// TIA Portal project "Project2_Pompe" (V15.1)

(* hardware
DEVICE "S71500/ET200MP station_1"  S7-1500 station
   slot 0: "Rail_0"  Rack  6ES7 590-1***0-0AA0
   slot 1: "PLC_1"  CPU 1513-1 PN  6ES7 513-1AL02-0AB0  V2.6
      slot 3: "CPU display_1"  6ES7591-1AA00-0AA0
DEVICE "HMI_1"  KTP900 Basic PN
   slot 0: "HMI_1"  KTP900 Basic PN  6AV2 123-2JB03-0AX0  15.1.0.0
   slot 1: "HMI_RT_1"  KTP900 Basic PN  6AV2 123-2JB03-0AX0  15.1.0.0
   slot 5: "HMI_1.IE_CP_1"  PROFINET Interface  15.0.1.0
      slot 1: "PROFINET Interface_1"  PROFINET Interface
         slot 1: "Port_1"  Port
*)

// ===== PLC "PLC_1"  CPU 1513-1 PN =====

VAR_GLOBAL   // PLC tag table "Default tag table"
   "Clock_Byte" AT %MB0 : Byte;
   "Clock_10Hz" AT %M0.0 : Bool;
   "Clock_5Hz" AT %M0.1 : Bool;
   "Clock_2.5Hz" AT %M0.2 : Bool;
   "Clock_2Hz" AT %M0.3 : Bool;
   "Clock_1.25Hz" AT %M0.4 : Bool;
   "Clock_1Hz" AT %M0.5 : Bool;
   "Clock_0.625Hz" AT %M0.6 : Bool;
   "Clock_0.5Hz" AT %M0.7 : Bool;
END_VAR

VAR_GLOBAL   // PLC tag table "Motor1"
   "permisie_start_1" AT %I0.0 : Bool;
   "motor_pornit_1" AT %I0.1 : Bool;
   "temporizare_k4_1" AT %I0.2 : Bool;
   "urgenta_bit_1" AT %I0.4 : Bool;
   "s1_1" AT %I0.7 : Bool;
   "s2_1" AT %I1.0 : Bool;
   "stop1" AT %I1.1 : Bool;
   "ptc1" AT %I1.2 : Bool;
   "timp_oprire_1" AT %ID1 : Time;
   "k1_1" AT %M1.4 : Bool;
   "k2_1" AT %M1.5 : Bool;
   "k3_1" AT %M1.6 : Bool;
   "k4_1" AT %M1.7 : Bool;
   "reset_urgenta_1" AT %I7.0 : Bool;
   "et_k4_1" AT %ID11 : Time;
   "et_stop_1" AT %ID10 : Time;
   "inactiv_1" AT %ID20 : Time;
END_VAR

VAR_GLOBAL   // PLC tag table "Motor2"
   "permisie_start_2" AT %I2.0 : Bool;
   "motor_pornit_2" AT %I2.1 : Bool;
   "temporizare_k4_2" AT %I2.2 : Bool;
   "urgenta_bit_2" AT %I2.3 : Bool;
   "s1_2" AT %I2.4 : Bool;
   "s2_2" AT %I2.5 : Bool;
   "stop2" AT %I2.6 : Bool;
   "ptc2" AT %I2.7 : Bool;
   "timp_oprire_2" AT %ID3 : Time;
   "k1_2" AT %M3.1 : Bool;
   "k2_2" AT %M3.2 : Bool;
   "k3_2" AT %M3.3 : Bool;
   "k4_2" AT %M3.4 : Bool;
   "reset_urgenta_2" AT %I7.1 : Bool;
   "et_k4_2" AT %ID7 : Time;
   "et_stop_2" AT %ID12 : Time;
   "inactiv_2" AT %ID16 : Time;
END_VAR

VAR_GLOBAL   // PLC tag table "Ambele_motoare"
   "ss(esd)" AT %I0.6 : Bool;
   "ptc" AT %I36.0 : Bool;
   "stop" AT %I36.1 : Bool;
   "reset_urgenta_general" AT %I36.2 : Bool;
   "urgenta_bit_ciuperca" AT %I36.3 : Bool;
   "oprire_toate_motoarele_pt_ptc" AT %I36.4 : Bool;
END_VAR

VAR_GLOBAL   // PLC tag table "Motor3"
   "permisie_start_3" AT %I30.0 : Bool;
   "motor_pornit_3" AT %I30.1 : Bool;
   "temporizare_k4_3" AT %I30.2 : Bool;
   "urgenta_bit_3" AT %I30.3 : Bool;
   "s1_3" AT %I30.4 : Bool;
   "s2_3" AT %I30.5 : Bool;
   "stop3" AT %I30.6 : Bool;
   "ptc3" AT %I30.7 : Bool;
   "k1_3" AT %M31.0 : Bool;
   "k2_3" AT %M31.1 : Bool;
   "k3_3" AT %M31.2 : Bool;
   "k4_3" AT %M31.3 : Bool;
   "reset_urgenta_3" AT %I31.4 : Bool;
   "et_k4_3" AT %ID31 : Time;
   "et_stop_3" AT %ID32 : Time;
END_VAR

VAR_GLOBAL   // PLC tag table "Motor4"
   "permisie_start_4" AT %I0.3 : Bool;
   "motor_pornit_4" AT %I0.5 : Bool;
   "temporizare_k4_4" AT %I24.0 : Bool;
   "urgenta_bit_4" AT %I24.1 : Bool;
   "s1_4" AT %I24.2 : Bool;
   "s2_4" AT %I24.3 : Bool;
   "stop4" AT %I24.4 : Bool;
   "pct4" AT %I24.5 : Bool;
   "k1_4" AT %M24.6 : Bool;
   "k2_4" AT %M24.7 : Bool;
   "k3_4" AT %M25.0 : Bool;
   "k4_4" AT %M25.1 : Bool;
   "reset_urgenta_4" AT %I25.2 : Bool;
   "et_k4_4" AT %ID25 : Time;
   "et_stop_4" AT %ID26 : Time;
END_VAR

DATA_BLOCK "db_directie_mers"   // DB1
{ S7_Optimized_Access := 'TRUE' }
VERSION : 0.1
   VAR
      et_stop : Time;
      stanga : Bool;
      dreapta : Bool;
      inainte : Bool;
      inapoi : Bool;
      stop : Bool;
   END_VAR
BEGIN
END_DATA_BLOCK

DATA_BLOCK "roata 2"   // DB3
{ S7_Optimized_Access := 'TRUE' }
VERSION : 0.1
// stored: InstanceOfName Fct_Motor
"Fct_Motor"
BEGIN
END_DATA_BLOCK

DATA_BLOCK "roata 3"   // DB4
{ S7_Optimized_Access := 'TRUE' }
VERSION : 0.1
// stored: InstanceOfName Fct_Motor
"Fct_Motor"
BEGIN
END_DATA_BLOCK

DATA_BLOCK "Alarme"   // DB5
{ S7_Optimized_Access := 'TRUE' }
VERSION : 0.1
   VAR
      alarme : Array[0..15] of Bool;
      alarme_merged : Word;
   END_VAR
BEGIN
END_DATA_BLOCK

DATA_BLOCK "functie ptc_DB_r1"   // DB7
{ S7_Optimized_Access := 'TRUE' }
VERSION : 0.1
// stored: InstanceOfName functie ptc
"functie ptc"
BEGIN
END_DATA_BLOCK

DATA_BLOCK "roata1"   // DB8
{ S7_Optimized_Access := 'TRUE' }
VERSION : 0.1
// stored: InstanceOfName Fct_Motor
"Fct_Motor"
BEGIN
END_DATA_BLOCK

DATA_BLOCK "roata 4"   // DB9
{ S7_Optimized_Access := 'TRUE' }
VERSION : 0.1
// stored: InstanceOfName Fct_Motor
"Fct_Motor"
BEGIN
END_DATA_BLOCK

DATA_BLOCK "functie ptc_DB_r2"   // DB10
{ S7_Optimized_Access := 'TRUE' }
VERSION : 0.1
// stored: InstanceOfName functie ptc
"functie ptc"
BEGIN
END_DATA_BLOCK

DATA_BLOCK "functie ptc_DB_r3"   // DB11
{ S7_Optimized_Access := 'TRUE' }
VERSION : 0.1
// stored: InstanceOfName functie ptc
"functie ptc"
BEGIN
END_DATA_BLOCK

DATA_BLOCK "functie ptc_DB_r4"   // DB12
{ S7_Optimized_Access := 'TRUE' }
VERSION : 0.1
// stored: InstanceOfName functie ptc
"functie ptc"
BEGIN
END_DATA_BLOCK

DATA_BLOCK "Data_block_1"   // DB13
{ S7_Optimized_Access := 'TRUE' }
VERSION : 0.1
   VAR
      tret : Bool;
      tret_1 : Bool;
      tret_2 : Bool;
      tret_3 : Bool;
      tret_4 : Bool;
      tret_5 : Bool;
      tret_6 : Bool;
   END_VAR
BEGIN
END_DATA_BLOCK

// folder: System blocks/Program resources

DATA_BLOCK "temp"   // DB2
{ S7_Optimized_Access := 'TRUE' }
AUTHOR : Simatic
FAMILY : IEC
NAME : IEC_TMR
VERSION : 1.0
// stored: InstanceOfName IEC_TIMER
"IEC_TIMER"
BEGIN
END_DATA_BLOCK

DATA_BLOCK "temp2"   // DB6
{ S7_Optimized_Access := 'TRUE' }
AUTHOR : Simatic
FAMILY : IEC
NAME : IEC_TMR
VERSION : 1.0
// stored: InstanceOfName IEC_TIMER
"IEC_TIMER"
BEGIN
END_DATA_BLOCK

// folder: (top level)

FUNCTION_BLOCK "Fct_Motor"   // FB1, LAD
{ S7_Optimized_Access := 'TRUE' }
VERSION : 0.1
   VAR_OUTPUT
      k1 : Bool;
      k2 : Bool;
      k3 : Bool;
      k4 : Bool;
   END_VAR
   VAR_IN_OUT
      "permisie start" : Bool;
      "motor pornit" : Bool;
      "temporizare k4" : Bool;
      "reset urgenta" : Bool;
      "urgenta bit" : Bool;
      s1 : Bool;
      s2 : Bool;
      ss : Bool;
      stop : Bool;
      ptc : Bool;
      et_stop : Time := T#0s;
      et_k4 : Time := T#0s;
   END_VAR
   VAR
      timerK4 : TON_TIME;
      timer_stop : TON_TIME;
   END_VAR
BEGIN

REGION Network 1: selecteaza k1
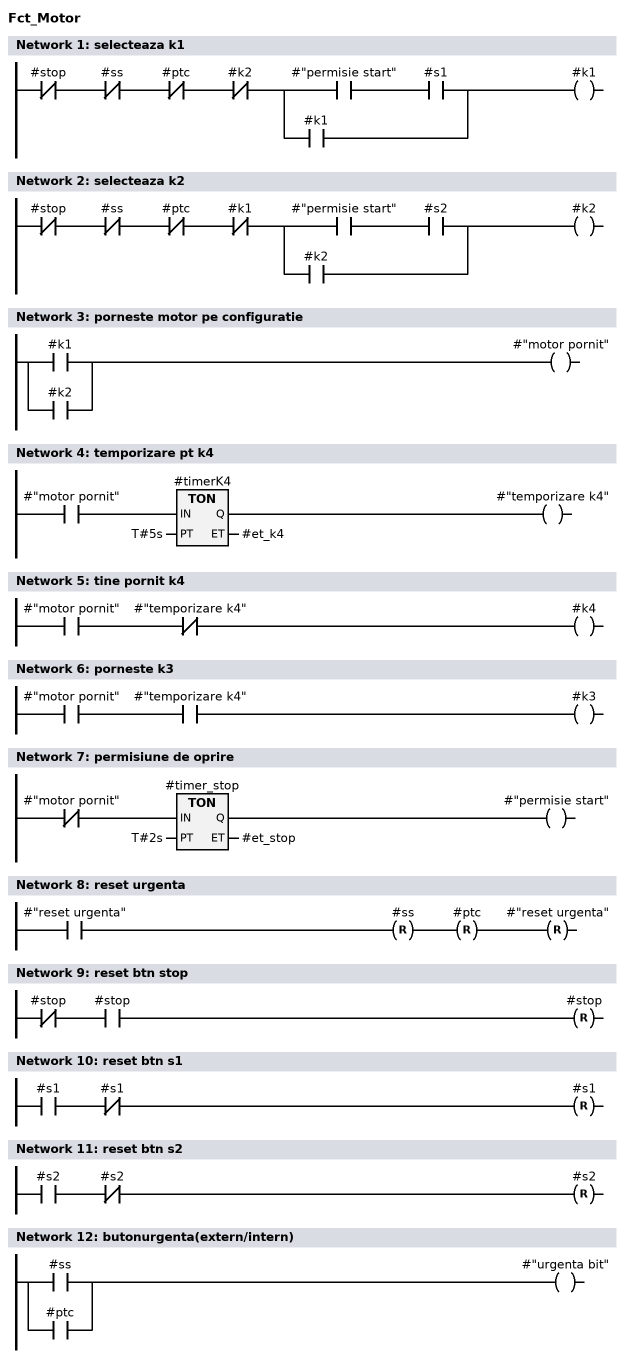
   RUNG wire#powerrail
      I_Contact( #stop )
      I_Contact( #ss )
      I_Contact( #ptc )
      I_Contact( #k2 )
      wire#w1
      Contact( #"permisie start" )
      Contact( #s1 )
      wire#w2
      Coil( #k1 )
   END_RUNG
   RUNG wire#w1
      Contact( #k1 )
   END_RUNG wire#w2
   // the same network as SCL:
   #k1 := NOT #stop AND NOT #ss AND NOT #ptc AND NOT #k2 AND ((#"permisie start" AND #s1) OR #k1);
END_REGION

REGION Network 2: selecteaza k2
   RUNG wire#powerrail
      I_Contact( #stop )
      I_Contact( #ss )
      I_Contact( #ptc )
      I_Contact( #k1 )
      wire#w1
      Contact( #"permisie start" )
      Contact( #s2 )
      wire#w2
      Coil( #k2 )
   END_RUNG
   RUNG wire#w1
      Contact( #k2 )
   END_RUNG wire#w2
   // the same network as SCL:
   #k2 := NOT #stop AND NOT #ss AND NOT #ptc AND NOT #k1 AND ((#"permisie start" AND #s2) OR #k2);
END_REGION

REGION Network 3: porneste motor pe configuratie
   RUNG wire#powerrail
      Contact( #k1 )
      wire#w1
      Coil( #"motor pornit" )
   END_RUNG
   RUNG wire#powerrail
      Contact( #k2 )
   END_RUNG wire#w1
   // the same network as SCL:
   #"motor pornit" := #k1 OR #k2;
END_REGION

REGION Network 4: temporizare pt k4
   #timerK4(IN := #"motor pornit", PT := T#5s, ET => #et_k4);   // TON
   #"temporizare k4" := #timerK4.Q;
END_REGION

REGION Network 5: tine pornit k4
   RUNG wire#powerrail
      Contact( #"motor pornit" )
      I_Contact( #"temporizare k4" )
      Coil( #k4 )
   END_RUNG
   // the same network as SCL:
   #k4 := #"motor pornit" AND NOT #"temporizare k4";
END_REGION

REGION Network 6: porneste k3
   RUNG wire#powerrail
      Contact( #"motor pornit" )
      Contact( #"temporizare k4" )
      Coil( #k3 )
   END_RUNG
   // the same network as SCL:
   #k3 := #"motor pornit" AND #"temporizare k4";
END_REGION

REGION Network 7: permisiune de oprire
   #timer_stop(IN := NOT #"motor pornit", PT := T#2s, ET => #et_stop);   // TON
   #"permisie start" := #timer_stop.Q;
END_REGION

REGION Network 8: reset urgenta
   RUNG wire#powerrail
      Contact( #"reset urgenta" )
      R_Coil( #ss )
      R_Coil( #ptc )
      R_Coil( #"reset urgenta" )
   END_RUNG
   // the same network as SCL:
   IF #"reset urgenta" THEN
       #ss := FALSE;
       #ptc := FALSE;
       #"reset urgenta" := FALSE;
   END_IF;
END_REGION

REGION Network 9: reset btn stop
   RUNG wire#powerrail
      I_Contact( #stop )
      Contact( #stop )
      R_Coil( #stop )
   END_RUNG
   // the same network as SCL:
   IF NOT #stop AND #stop THEN #stop := FALSE; END_IF;
END_REGION

REGION Network 10: reset btn s1
   RUNG wire#powerrail
      Contact( #s1 )
      I_Contact( #s1 )
      R_Coil( #s1 )
   END_RUNG
   // the same network as SCL:
   IF #s1 AND NOT #s1 THEN #s1 := FALSE; END_IF;
END_REGION

REGION Network 11: reset btn s2
   RUNG wire#powerrail
      Contact( #s2 )
      I_Contact( #s2 )
      R_Coil( #s2 )
   END_RUNG
   // the same network as SCL:
   IF #s2 AND NOT #s2 THEN #s2 := FALSE; END_IF;
END_REGION

REGION Network 12: butonurgenta(extern/intern)
   RUNG wire#powerrail
      Contact( #ss )
      wire#w1
      Coil( #"urgenta bit" )
   END_RUNG
   RUNG wire#powerrail
      Contact( #ptc )
   END_RUNG wire#w1
   // the same network as SCL:
   #"urgenta bit" := #ss OR #ptc;
END_REGION
END_FUNCTION_BLOCK

FUNCTION_BLOCK "functie ptc"   // FB2, LAD
{ S7_Optimized_Access := 'TRUE' }
VERSION : 0.1
   VAR_OUTPUT
      alarma : Bool;
   END_VAR
   VAR_IN_OUT
      reset_urgenta : Bool;
      ptc_apasat : Bool;
   END_VAR
   VAR
      timer_buton_reset : TON_TIME;
      IEC_Timer_0_Instance : TON_TIME;
   END_VAR
BEGIN

REGION Network 1: apasa butonul
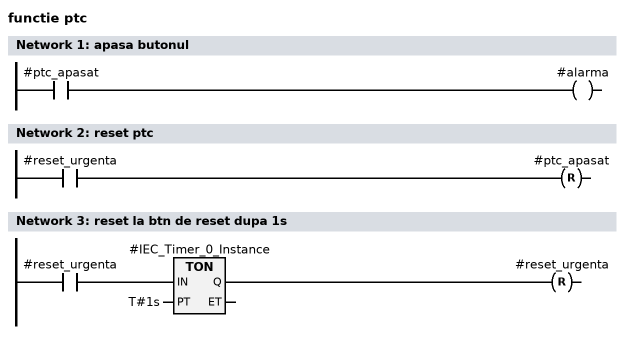
   RUNG wire#powerrail
      Contact( #ptc_apasat )
      Coil( #alarma )
   END_RUNG
   // the same network as SCL:
   #alarma := #ptc_apasat;
END_REGION

REGION Network 2: reset ptc
   RUNG wire#powerrail
      Contact( #reset_urgenta )
      R_Coil( #ptc_apasat )
   END_RUNG
   // the same network as SCL:
   IF #reset_urgenta THEN #ptc_apasat := FALSE; END_IF;
END_REGION

REGION Network 3: reset la btn de reset dupa 1s
   #IEC_Timer_0_Instance(IN := #reset_urgenta, PT := T#1s);   // TON
   IF #IEC_Timer_0_Instance.Q THEN #reset_urgenta := FALSE; END_IF;
END_REGION
END_FUNCTION_BLOCK

ORGANIZATION_BLOCK "Main"   // OB1, LAD, ProgramCycle
TITLE = "Main Program Sweep (Cycle)"
{ S7_Optimized_Access := 'TRUE' }
VERSION : 0.1
   VAR_INPUT
      Initial_Call : Bool;   // Initial call of this OB
      Remanence : Bool;   // =True, if remanent data are available
   END_VAR
   VAR_TEMP   // added for the SCL form of the ladder/FBD networks
      _w1 : Bool;
      _w2 : Bool;
      _w3 : Bool;
   END_VAR
BEGIN

REGION Network 1: initializare cele 2 roti fata
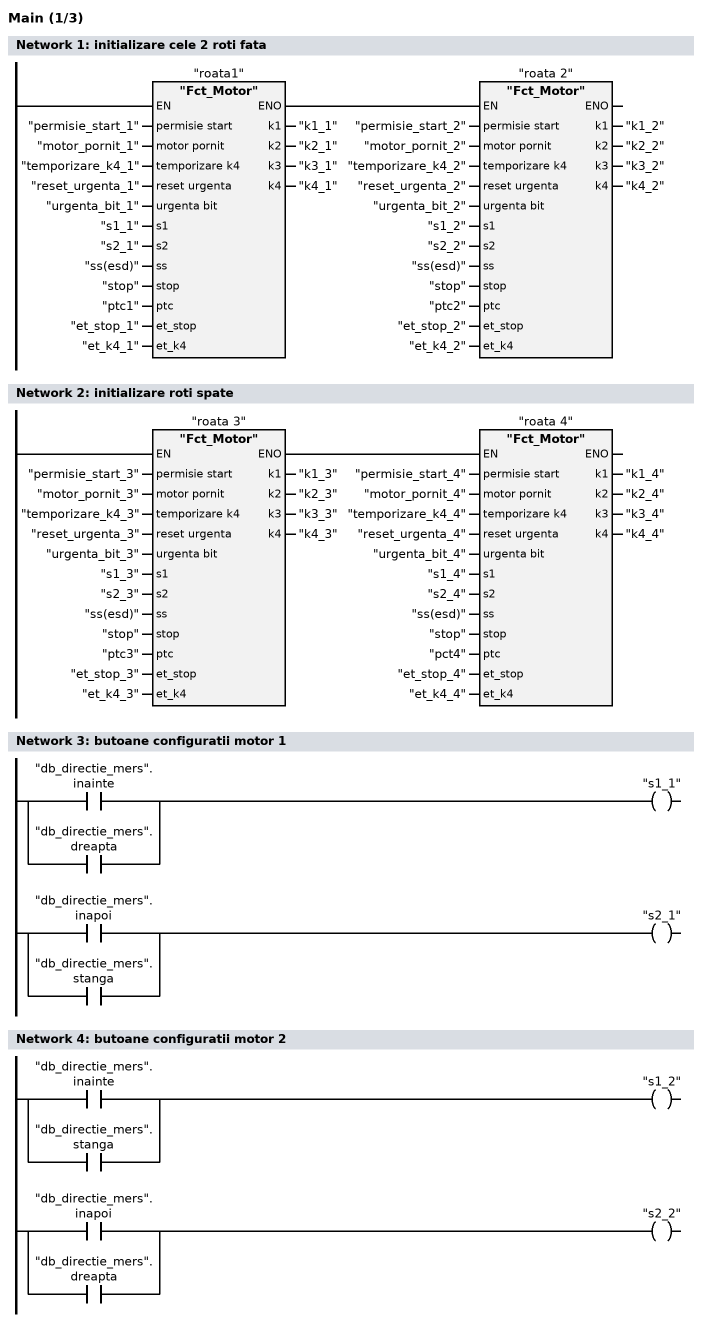
   RUNG wire#powerrail
      "roata1"("permisie start" := "permisie_start_1", "motor pornit" := "motor_pornit_1", "temporizare k4" := "temporizare_k4_1", "reset urgenta" := "reset_urgenta_1", "urgenta bit" := "urgenta_bit_1", s1 := "s1_1", s2 := "s2_1", ss := "ss(esd)", stop := "stop", ptc := "ptc1", et_stop := "et_stop_1", et_k4 := "et_k4_1", k1 => "k1_1", k2 => "k2_1", k3 => "k3_1", k4 => "k4_1")
      "roata 2"("permisie start" := "permisie_start_2", "motor pornit" := "motor_pornit_2", "temporizare k4" := "temporizare_k4_2", "reset urgenta" := "reset_urgenta_2", "urgenta bit" := "urgenta_bit_2", s1 := "s1_2", s2 := "s2_2", ss := "ss(esd)", stop := "stop", ptc := "ptc2", et_stop := "et_stop_2", et_k4 := "et_k4_2", k1 => "k1_2", k2 => "k2_2", k3 => "k3_2", k4 => "k4_2")
   END_RUNG
   // the same network as SCL:
   "roata1"("permisie start" := "permisie_start_1",   // "Fct_Motor"
            "motor pornit" := "motor_pornit_1",
            "temporizare k4" := "temporizare_k4_1",
            "reset urgenta" := "reset_urgenta_1",
            "urgenta bit" := "urgenta_bit_1",
            s1 := "s1_1",
            s2 := "s2_1",
            ss := "ss(esd)",
            stop := "stop",
            ptc := "ptc1",
            et_stop := "et_stop_1",
            et_k4 := "et_k4_1",
            k1 => "k1_1",
            k2 => "k2_1",
            k3 => "k3_1",
            k4 => "k4_1",
            ENO => #_w1);
   IF #_w1 THEN
       "roata 2"("permisie start" := "permisie_start_2",   // "Fct_Motor"
                 "motor pornit" := "motor_pornit_2",
                 "temporizare k4" := "temporizare_k4_2",
                 "reset urgenta" := "reset_urgenta_2",
                 "urgenta bit" := "urgenta_bit_2",
                 s1 := "s1_2",
                 s2 := "s2_2",
                 ss := "ss(esd)",
                 stop := "stop",
                 ptc := "ptc2",
                 et_stop := "et_stop_2",
                 et_k4 := "et_k4_2",
                 k1 => "k1_2",
                 k2 => "k2_2",
                 k3 => "k3_2",
                 k4 => "k4_2");
   END_IF;
END_REGION

REGION Network 2: initializare roti spate
   RUNG wire#powerrail
      "roata 3"("permisie start" := "permisie_start_3", "motor pornit" := "motor_pornit_3", "temporizare k4" := "temporizare_k4_3", "reset urgenta" := "reset_urgenta_3", "urgenta bit" := "urgenta_bit_3", s1 := "s1_3", s2 := "s2_3", ss := "ss(esd)", stop := "stop", ptc := "ptc3", et_stop := "et_stop_3", et_k4 := "et_k4_3", k1 => "k1_3", k2 => "k2_3", k3 => "k3_3", k4 => "k4_3")
      "roata 4"("permisie start" := "permisie_start_4", "motor pornit" := "motor_pornit_4", "temporizare k4" := "temporizare_k4_4", "reset urgenta" := "reset_urgenta_4", "urgenta bit" := "urgenta_bit_4", s1 := "s1_4", s2 := "s2_4", ss := "ss(esd)", stop := "stop", ptc := "pct4", et_stop := "et_stop_4", et_k4 := "et_k4_4", k1 => "k1_4", k2 => "k2_4", k3 => "k3_4", k4 => "k4_4")
   END_RUNG
   // the same network as SCL:
   "roata 3"("permisie start" := "permisie_start_3",   // "Fct_Motor"
             "motor pornit" := "motor_pornit_3",
             "temporizare k4" := "temporizare_k4_3",
             "reset urgenta" := "reset_urgenta_3",
             "urgenta bit" := "urgenta_bit_3",
             s1 := "s1_3",
             s2 := "s2_3",
             ss := "ss(esd)",
             stop := "stop",
             ptc := "ptc3",
             et_stop := "et_stop_3",
             et_k4 := "et_k4_3",
             k1 => "k1_3",
             k2 => "k2_3",
             k3 => "k3_3",
             k4 => "k4_3",
             ENO => #_w1);
   IF #_w1 THEN
       "roata 4"("permisie start" := "permisie_start_4",   // "Fct_Motor"
                 "motor pornit" := "motor_pornit_4",
                 "temporizare k4" := "temporizare_k4_4",
                 "reset urgenta" := "reset_urgenta_4",
                 "urgenta bit" := "urgenta_bit_4",
                 s1 := "s1_4",
                 s2 := "s2_4",
                 ss := "ss(esd)",
                 stop := "stop",
                 ptc := "pct4",
                 et_stop := "et_stop_4",
                 et_k4 := "et_k4_4",
                 k1 => "k1_4",
                 k2 => "k2_4",
                 k3 => "k3_4",
                 k4 => "k4_4");
   END_IF;
END_REGION

REGION Network 3: butoane configuratii motor 1
   RUNG wire#powerrail
      Contact( "db_directie_mers".inainte )
      wire#w1
      Coil( "s1_1" )
   END_RUNG
   RUNG wire#powerrail
      Contact( "db_directie_mers".dreapta )
   END_RUNG wire#w1
   RUNG wire#powerrail
      Contact( "db_directie_mers".inapoi )
      wire#w2
      Coil( "s2_1" )
   END_RUNG
   RUNG wire#powerrail
      Contact( "db_directie_mers".stanga )
   END_RUNG wire#w2
   // the same network as SCL:
   "s1_1" := "db_directie_mers".inainte OR "db_directie_mers".dreapta;
   "s2_1" := "db_directie_mers".inapoi OR "db_directie_mers".stanga;
END_REGION

REGION Network 4: butoane configuratii motor 2
   RUNG wire#powerrail
      Contact( "db_directie_mers".inainte )
      wire#w1
      Coil( "s1_2" )
   END_RUNG
   RUNG wire#powerrail
      Contact( "db_directie_mers".stanga )
   END_RUNG wire#w1
   RUNG wire#powerrail
      Contact( "db_directie_mers".inapoi )
      wire#w2
      Coil( "s2_2" )
   END_RUNG
   RUNG wire#powerrail
      Contact( "db_directie_mers".dreapta )
   END_RUNG wire#w2
   // the same network as SCL:
   "s1_2" := "db_directie_mers".inainte OR "db_directie_mers".stanga;
   "s2_2" := "db_directie_mers".inapoi OR "db_directie_mers".dreapta;
END_REGION

REGION Network 5: butoane configuratii motor 3
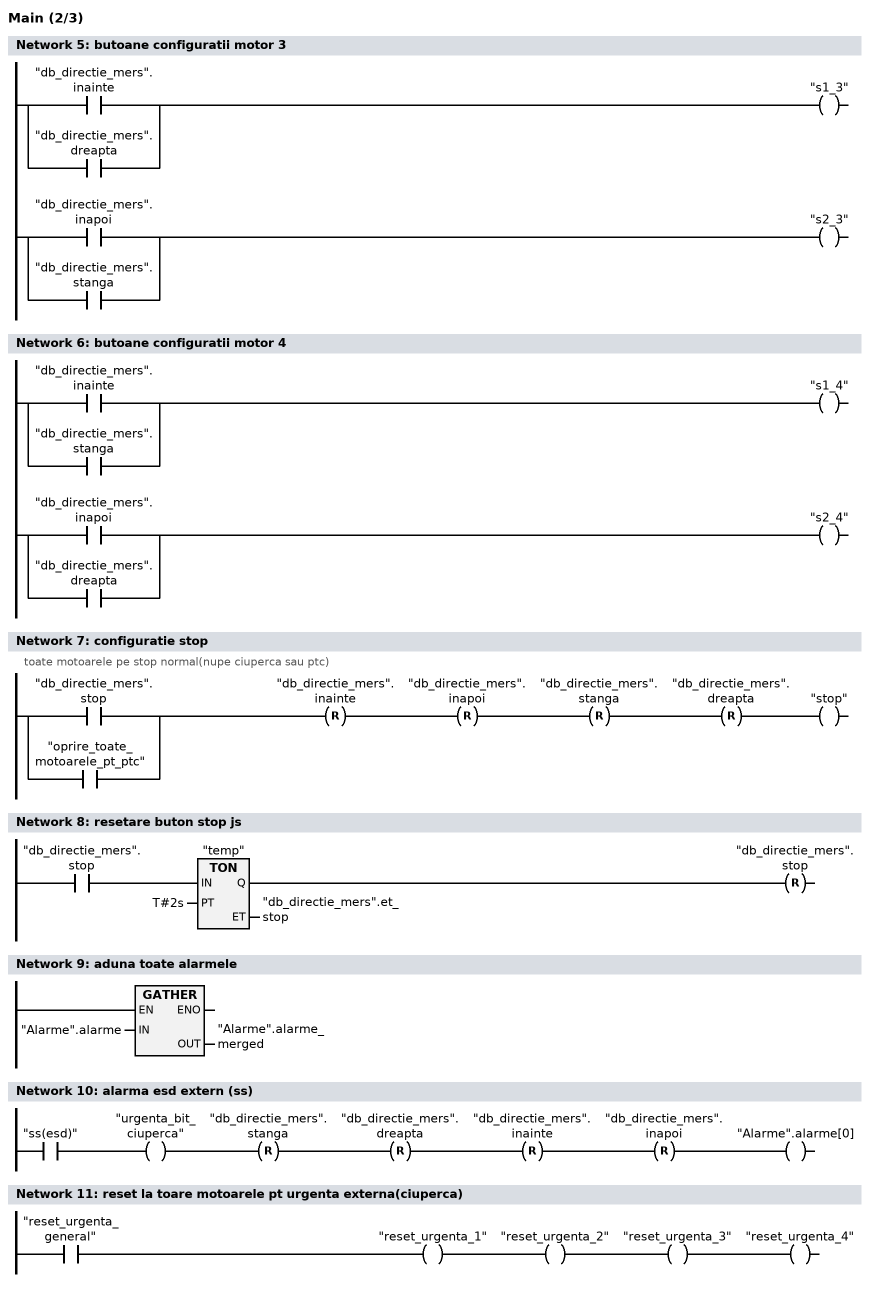
   RUNG wire#powerrail
      Contact( "db_directie_mers".inainte )
      wire#w1
      Coil( "s1_3" )
   END_RUNG
   RUNG wire#powerrail
      Contact( "db_directie_mers".dreapta )
   END_RUNG wire#w1
   RUNG wire#powerrail
      Contact( "db_directie_mers".inapoi )
      wire#w2
      Coil( "s2_3" )
   END_RUNG
   RUNG wire#powerrail
      Contact( "db_directie_mers".stanga )
   END_RUNG wire#w2
   // the same network as SCL:
   "s1_3" := "db_directie_mers".inainte OR "db_directie_mers".dreapta;
   "s2_3" := "db_directie_mers".inapoi OR "db_directie_mers".stanga;
END_REGION

REGION Network 6: butoane configuratii motor 4
   RUNG wire#powerrail
      Contact( "db_directie_mers".inainte )
      wire#w1
      Coil( "s1_4" )
   END_RUNG
   RUNG wire#powerrail
      Contact( "db_directie_mers".stanga )
   END_RUNG wire#w1
   RUNG wire#powerrail
      Contact( "db_directie_mers".inapoi )
      wire#w2
      Coil( "s2_4" )
   END_RUNG
   RUNG wire#powerrail
      Contact( "db_directie_mers".dreapta )
   END_RUNG wire#w2
   // the same network as SCL:
   "s1_4" := "db_directie_mers".inainte OR "db_directie_mers".stanga;
   "s2_4" := "db_directie_mers".inapoi OR "db_directie_mers".dreapta;
END_REGION

REGION Network 7: configuratie stop
   // toate motoarele pe stop normal(nupe ciuperca sau ptc)
   RUNG wire#powerrail
      Contact( "db_directie_mers".stop )
      wire#w1
      R_Coil( "db_directie_mers".inainte )
      R_Coil( "db_directie_mers".inapoi )
      R_Coil( "db_directie_mers".stanga )
      R_Coil( "db_directie_mers".dreapta )
      Coil( "stop" )
   END_RUNG
   RUNG wire#powerrail
      Contact( "oprire_toate_motoarele_pt_ptc" )
   END_RUNG wire#w1
   // the same network as SCL:
   #_w1 := "db_directie_mers".stop OR "oprire_toate_motoarele_pt_ptc";
   IF #_w1 THEN
       "db_directie_mers".inainte := FALSE;
       "db_directie_mers".inapoi := FALSE;
       "db_directie_mers".stanga := FALSE;
       "db_directie_mers".dreapta := FALSE;
   END_IF;
   "stop" := #_w1;
END_REGION

REGION Network 8: resetare buton stop js
   "temp".TON(IN := "db_directie_mers".stop, PT := T#2s, ET => "db_directie_mers".et_stop);
   IF "temp".Q THEN "db_directie_mers".stop := FALSE; END_IF;
END_REGION

REGION Network 9: aduna toate alarmele
   GATHER(IN := "Alarme".alarme, OUT => "Alarme".alarme_merged);
END_REGION

REGION Network 10: alarma esd extern (ss)
   RUNG wire#powerrail
      Contact( "ss(esd)" )
      Coil( "urgenta_bit_ciuperca" )
      R_Coil( "db_directie_mers".stanga )
      R_Coil( "db_directie_mers".dreapta )
      R_Coil( "db_directie_mers".inainte )
      R_Coil( "db_directie_mers".inapoi )
      Coil( "Alarme".alarme[0] )
   END_RUNG
   // the same network as SCL:
   "urgenta_bit_ciuperca" := "ss(esd)";
   IF "ss(esd)" THEN
       "db_directie_mers".stanga := FALSE;
       "db_directie_mers".dreapta := FALSE;
       "db_directie_mers".inainte := FALSE;
       "db_directie_mers".inapoi := FALSE;
   END_IF;
   "Alarme".alarme[0] := "ss(esd)";
END_REGION

REGION Network 11: reset la toare motoarele pt urgenta externa(ciuperca)
   RUNG wire#powerrail
      Contact( "reset_urgenta_general" )
      Coil( "reset_urgenta_1" )
      Coil( "reset_urgenta_2" )
      Coil( "reset_urgenta_3" )
      Coil( "reset_urgenta_4" )
   END_RUNG
   // the same network as SCL:
   "reset_urgenta_1" := "reset_urgenta_general";
   "reset_urgenta_2" := "reset_urgenta_general";
   "reset_urgenta_3" := "reset_urgenta_general";
   "reset_urgenta_4" := "reset_urgenta_general";
END_REGION

REGION Network 12: reset la butonul de reset general dupa 1s
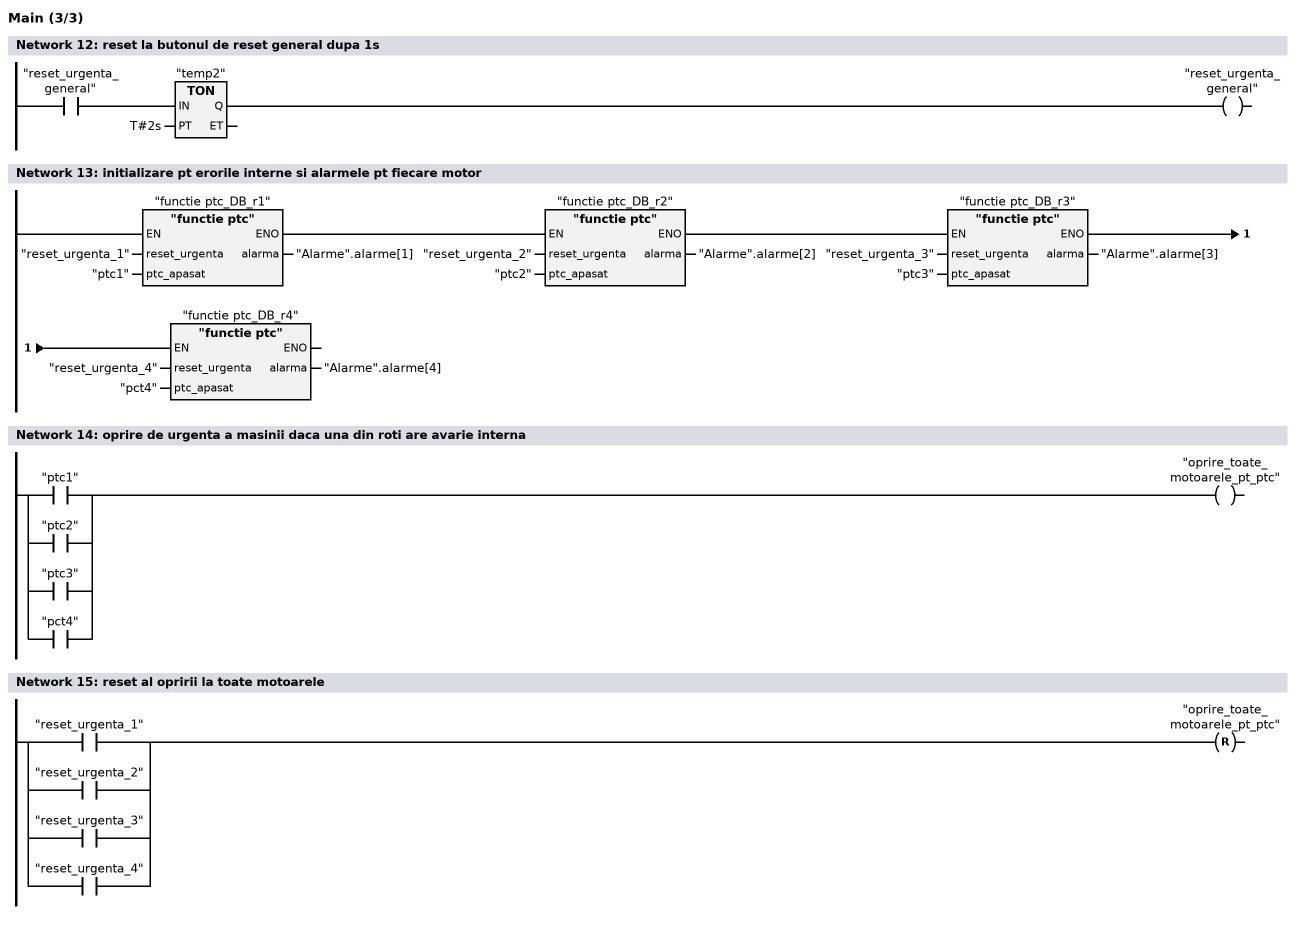
   "temp2".TON(IN := "reset_urgenta_general", PT := T#2s);
   "reset_urgenta_general" := "temp2".Q;
END_REGION

REGION Network 13: initializare pt erorile interne si alarmele pt fiecare motor
   RUNG wire#powerrail
      "functie ptc_DB_r1"(reset_urgenta := "reset_urgenta_1", ptc_apasat := "ptc1", alarma => "Alarme".alarme[1])
      "functie ptc_DB_r2"(reset_urgenta := "reset_urgenta_2", ptc_apasat := "ptc2", alarma => "Alarme".alarme[2])
      "functie ptc_DB_r3"(reset_urgenta := "reset_urgenta_3", ptc_apasat := "ptc3", alarma => "Alarme".alarme[3])
      "functie ptc_DB_r4"(reset_urgenta := "reset_urgenta_4", ptc_apasat := "pct4", alarma => "Alarme".alarme[4])
   END_RUNG
   // the same network as SCL:
   "functie ptc_DB_r1"(reset_urgenta := "reset_urgenta_1",   // "functie ptc"
                       ptc_apasat := "ptc1",
                       alarma => "Alarme".alarme[1],
                       ENO => #_w1);
   "functie ptc_DB_r2"(EN := #_w1,   // "functie ptc"
                       reset_urgenta := "reset_urgenta_2",
                       ptc_apasat := "ptc2",
                       alarma => "Alarme".alarme[2],
                       ENO => #_w2);
   "functie ptc_DB_r3"(EN := #_w2,   // "functie ptc"
                       reset_urgenta := "reset_urgenta_3",
                       ptc_apasat := "ptc3",
                       alarma => "Alarme".alarme[3],
                       ENO => #_w3);
   IF #_w3 THEN
       "functie ptc_DB_r4"(reset_urgenta := "reset_urgenta_4", ptc_apasat := "pct4", alarma => "Alarme".alarme[4]);   // "functie ptc"
   END_IF;
END_REGION

REGION Network 14: oprire de urgenta a masinii daca una din roti are avarie interna
   RUNG wire#powerrail
      Contact( "ptc1" )
      wire#w1
      Coil( "oprire_toate_motoarele_pt_ptc" )
   END_RUNG
   RUNG wire#powerrail
      Contact( "ptc2" )
   END_RUNG wire#w1
   RUNG wire#powerrail
      Contact( "ptc3" )
   END_RUNG wire#w1
   RUNG wire#powerrail
      Contact( "pct4" )
   END_RUNG wire#w1
   // the same network as SCL:
   "oprire_toate_motoarele_pt_ptc" := "ptc1" OR "ptc2" OR "ptc3" OR "pct4";
END_REGION

REGION Network 15: reset al opririi la toate motoarele
   RUNG wire#powerrail
      Contact( "reset_urgenta_1" )
      wire#w1
      R_Coil( "oprire_toate_motoarele_pt_ptc" )
   END_RUNG
   RUNG wire#powerrail
      Contact( "reset_urgenta_2" )
   END_RUNG wire#w1
   RUNG wire#powerrail
      Contact( "reset_urgenta_3" )
   END_RUNG wire#w1
   RUNG wire#powerrail
      Contact( "reset_urgenta_4" )
   END_RUNG wire#w1
   // the same network as SCL:
   IF "reset_urgenta_1" OR "reset_urgenta_2" OR "reset_urgenta_3" OR "reset_urgenta_4" THEN
       "oprire_toate_motoarele_pt_ptc" := FALSE;
   END_IF;
END_REGION
END_ORGANIZATION_BLOCK

(* ===== HMI "HMI_RT_1" =====
system functions are stored by id; their names below are inferred from use
connection "HMI_Connection_1": ETHERNET, SMART_S7_1500_OMS

HMI tags "Default tag table"
   "stop1" : Bool = PLC stop1 AT %I1.1, 1 s
   "s1_1" : Bool = PLC s1_1 AT %I0.7, 1 s
   "s2_1" : Bool = PLC s2_1 AT %I1.0, 1 s
   "k1_1" : Bool = PLC k1_1 AT %M1.4, 1 s
   "k2_1" : Bool = PLC k2_1 AT %M1.5, 1 s
   "urgenta_bit_1" : Bool = PLC urgenta_bit_1 AT %I0.4, 1 s
   "ptc1" : Bool = PLC ptc1 AT %I1.2, 1 s
   "k4_1" : Bool = PLC k4_1 AT %M1.7, 1 s
   "k3_1" : Bool = PLC k3_1 AT %M1.6, 1 s
   "timp_oprire_1" : Time = PLC timp_oprire_1 AT %ID1, 1 s
   "motor_pornit_1" : Bool = PLC motor_pornit_1 AT %I0.1, 1 s
   "stop2" : Bool = PLC stop2 AT %I2.6, 1 s
   "s1_2" : Bool = PLC s1_2 AT %I2.4, 1 s
   "s2_2" : Bool = PLC s2_2 AT %I2.5, 1 s
   "k1_2" : Bool = PLC k1_2 AT %M3.1, 1 s
   "k2_2" : Bool = PLC k2_2 AT %M3.2, 1 s
   "urgenta_bit_2" : Bool = PLC urgenta_bit_2 AT %I2.3, 1 s
   "ptc2" : Bool = PLC ptc2 AT %I2.7, 1 s
   "reset_urgenta_1" : Bool = PLC reset_urgenta_1 AT %I7.0, 1 s
   "reset_urgenta_2" : Bool = PLC reset_urgenta_2 AT %I7.1, 1 s
   "k4_2" : Bool = PLC k4_2 AT %M3.4, 1 s
   "k3_2" : Bool = PLC k3_2 AT %M3.3, 1 s
   "motor_pornit_2" : Bool = PLC motor_pornit_2 AT %I2.1, 1 s
   "ss" : Bool = PLC "ss(esd)" AT %I0.6, 1 s
   "et_k4_1" : Time = PLC et_k4_1 AT %ID11, 1 s
   "et_stop_1" : Time = PLC et_stop_1 AT %ID10, 1 s
   "et_stop_2" : Time = PLC et_stop_2 AT %ID12, 1 s
   "et_k4_2" : Time = PLC et_k4_2 AT %ID7, 1 s
   "inactiv_2" : Time = PLC inactiv_2 AT %ID16, 1 s
   "inactiv_1" : Time = PLC inactiv_1 AT %ID20, 1 s
   "Data_block_1_alarme_merged" : Word = PLC Alarme.alarme_merged, 1 s
   "reset_urgenta_general" : Bool = PLC reset_urgenta_general AT %I36.2, 1 s
   "urgenta_bit_ciuperca" : Bool = PLC urgenta_bit_ciuperca AT %I36.3, 1 s
   "stop" : Bool = PLC stop AT %I36.1, 1 s
   "db_directie_mers_inainte" : Bool = PLC db_directie_mers.inainte, 1 s
   "db_directie_mers_stop" : Bool = PLC db_directie_mers.stop, 1 s
   "db_directie_mers_inapoi" : Bool = PLC db_directie_mers.inapoi, 1 s
   "db_directie_mers_stanga" : Bool = PLC db_directie_mers.stanga, 1 s
   "db_directie_mers_dreapta" : Bool = PLC db_directie_mers.dreapta, 1 s
   "k1_3" : Bool = PLC k1_3 AT %M31.0, 1 s
   "k2_3" : Bool = PLC k2_3 AT %M31.1, 1 s
   "k1_4" : Bool = PLC k1_4 AT %M24.6, 1 s
   "k2_4" : Bool = PLC k2_4 AT %M24.7, 1 s
   "db_directie_mers_et_stop" : Time = PLC db_directie_mers.et_stop, 1 s
   "ptc3" : Bool = PLC ptc3 AT %I30.7, 1 s
   "pct4" : Bool = PLC pct4 AT %I24.5, 1 s
   "reset_urgenta_3" : Bool = PLC reset_urgenta_3 AT %I31.4, 1 s
   "reset_urgenta_4" : Bool = PLC reset_urgenta_4 AT %I25.2, 1 s

discrete alarms
   1: 'S-a apasat ciuperca boss', class Errors, trigger "Data_block_1_alarme_merged" bit 0
   2: 'Motorul de la roata 1 nu mai merge', class Errors, trigger "Data_block_1_alarme_merged" bit 1
   3: 'Motorul de la roata 2 nu mai merge', class Errors, trigger "Data_block_1_alarme_merged" bit 2
   4: 'Motorul de la roata 3 nu mai merge', class Errors, trigger "Data_block_1_alarme_merged" bit 3
   5: 'Motorul de la roata 4 nu mai merge', class Errors, trigger "Data_block_1_alarme_merged" bit 4
   6: '', class Errors, trigger "Data_block_1_alarme_merged" bit 5
   7: '', class Errors, trigger "Data_block_1_alarme_merged" bit 6

Template "Template_1" 800x480
   Button "Exit" at 722,440 size 55x39; TextOff 'Exit'; PictureOff "ExitRuntime_KTP900_Basic_PN_TR"; PictureOn "ExitRuntime_KTP900_Basic_PN_TR"
      on Release: StopRuntime(0)
   Button "Template_Button" at 622,440 size 55x39; TextOff 'Text'
   Button "Template_Button_1" at 522,440 size 55x39; TextOff 'Text'
   Button "Template_Button_2" at 422,440 size 55x39; TextOff 'Text'
   Button "Template_Button_3" at 322,440 size 55x39; TextOff 'Text'
   Button "Template_Button_4" at 222,440 size 55x39; TextOff 'Text'
   Button "Alarms" at 122,440 size 55x39; TextOff 'Alarms'; PictureOff "AlarmDisplay_KTP900_Basic_PN_TR"; PictureOn "AlarmDisplay_KTP900_Basic_PN_TR"
      on Release: function_ef3f5d25("Alarm window_1", -1)
   Button "Start screen" at 22,440 size 55x39; TextOff 'Start screen'; PictureOff "NavigateHome_KTP900_Basic_PN_TR"; PictureOn "NavigateHome_KTP900_Basic_PN_TR"
      on Release: ActivateScreen("Root screen", 0)
   DateTimeField "HmiScreenItemData" at 695,20 size 105x20
   DateTimeField "HmiScreenItemData_1" at 695,0 size 105x20
   GraphicView "Logo" at 0,0 size 71x40; Picture "Logo of HMI_1"

screen "Root screen" 800x480, template "Template_1"
   Button "Button_4" at 623,351 size 96x32; TextOff 'ESD'
      on Click: SetBit("ss")
   TextField "Text field_7" at 584,353 size 21x20; Text 'SS'
   Button "Button_5" at 21,390 size 96x32; TextOff 'Just press'
   Button "Button_6" at 623,397 size 96x32; TextOff 'Reset ESD'
      on Click: SetBit("reset_urgenta_general")
   Ellipse "Ellipse_1" at 640,317 size 67x28
      Appearance <- "urgenta_bit_ciuperca"
   IOField "I/O field_2" at 231,378 size 96x32; FormatPattern 99999; Unit ms
      ProcessValue <- "et_stop_2"
   TextField "Text field_11" at 257,353 size 73x20; Text 'Timer stop'
   Button "Button_1" at 639,43 size 40x81; TextOff 'Fata'
      on Click: SetBit("db_directie_mers_inainte")
   Button "Button_2" at 640,185 size 42x81; TextOff 'Spate'
      on Click: SetBit("db_directie_mers_inapoi")
   Button "Button_3" at 527,143 size 96x32; TextOff 'Stanga'
      on Click: SetBit("db_directie_mers_stanga")
   Button "Button_7" at 698,143 size 96x32; TextOff 'Dreapta'
      on Click: SetBit("db_directie_mers_dreapta")
   Button "Button_8" at 637,141 size 49x32; TextOff 'Stop'
      on Click: SetBit("db_directie_mers_stop")
   TextField "Text field_1" at 298,31 size 89x20; Text 'Configuratie:'
   Button "Button_9" at 327,173 size 52x32; TextOff 'PTC1'
   Button "Button_10" at 387,173 size 36x32; TextOff 'R1'
   Button "Button_11" at 327,216 size 52x32; TextOff 'PTC2'
      on Click: SetBit("ptc2")
   Button "Button_12" at 387,216 size 36x32; TextOff 'R2'
      on Click: SetBit("reset_urgenta_2")
   Circle "Circle_3" at 436,216 size 30x30
      Appearance <- "ptc2"
   Button "Button_13" at 327,173 size 52x32; TextOff 'PTC1'
      on Click: SetBit("ptc1")
   Button "Button_14" at 387,173 size 36x32; TextOff 'R1'
      on Click: SetBit("reset_urgenta_1")
   Circle "Circle_4" at 436,173 size 30x30
      Appearance <- "ptc1"
   Button "Button_15" at 327,255 size 52x32; TextOff 'PTC3'
      on Click: SetBit("ptc3")
   Button "Button_16" at 387,255 size 36x32; TextOff 'R3'
      on Click: SetBit("reset_urgenta_3")
   Circle "Circle_5" at 436,255 size 30x30
      Appearance <- "ptc3"
   Button "Button_17" at 327,295 size 52x32; TextOff 'PTC4'
      on Click: SetBit("pct4")
   Button "Button_18" at 387,295 size 36x32; TextOff 'R4'
      on Click: SetBit("reset_urgenta_4")
   Circle "Circle_9" at 436,295 size 30x30
      Appearance <- "pct4"
   TextField "Text field_2" at 413,31 size 51x20; Text 'Inainte'
      Visibility <- "db_directie_mers_inainte"
   TextField "Text field_3" at 415,31 size 45x20; Text 'Inapoi'
      Visibility <- "db_directie_mers_inapoi"
   TextField "Text field_4" at 425,31 size 35x20; Text 'Stop'
      Visibility <- "db_directie_mers_stop"
   TextField "Text field_5" at 409,31 size 51x20; Text 'Stanga'
      Visibility <- "db_directie_mers_stanga"
   TextField "Text field_6" at 402,31 size 58x20; Text 'Dreapta'
      Visibility <- "db_directie_mers_dreapta"
   Rectangle "Rectangle_1" at 21,269 size 34x48
      Appearance <- "k1_3"
   Rectangle "Rectangle_2" at 54,269 size 34x48
      Appearance <- "k2_3"
   Rectangle "Rectangle_3" at 123,90 size 34x48
      Appearance <- "k1_2"
   Rectangle "Rectangle_4" at 156,90 size 34x48
      Appearance <- "k2_2"
   Rectangle "Rectangle_5" at 20,91 size 34x48
      Appearance <- "k1_1"
   Rectangle "Rectangle_6" at 53,91 size 34x48
      Appearance <- "k2_1"
   Rectangle "Rectangle_7" at 134,269 size 34x48
      Appearance <- "k1_4"
   Rectangle "Rectangle_8" at 167,269 size 34x48
      Appearance <- "k2_4"
   TextField "Text field_8" at 42,57 size 22x20; Text 'R1'
   TextField "Text field_9" at 146,57 size 22x20; Text 'R2'
   TextField "Text field_10" at 41,235 size 22x20; Text 'R3'
   TextField "Text field_12" at 159,235 size 22x20; Text 'R4'
   TextField "Text field_13" at 32,104 size 21x20; Text 'K1'
   TextField "Text field_14" at 141,285 size 21x20; Text 'K1'
   TextField "Text field_15" at 33,283 size 21x20; Text 'K1'
   TextField "Text field_16" at 134,100 size 21x20; Text 'K1'
   TextField "Text field_17" at 169,285 size 21x20; Text 'K2'
   TextField "Text field_18" at 159,100 size 21x20; Text 'K2'
   TextField "Text field_19" at 55,283 size 21x20; Text 'K2'
   TextField "Text field_25" at 54,104 size 21x20; Text 'K2'
*)